
screen "Nas_23" 1280x800
   Softkey "Softkey_F1" at 0,0 size 0x0
      on KeyDown: function_efd93a16()
   IOField "I/O field_6" at 38,288 size 172x31; FormatPattern s999.9; Unit %
      ProcessValue <- "PV"
   IOField "I/O field_1" at 35,197 size 174x31; FormatPattern s999.9; Unit %
      ProcessValue <- "SP"
   IOField "I/O field_2" at 240,288 size 149x31; FormatPattern s999.9; Unit %
      ProcessValue <- "LMN"
   TextField "Text field_8" at 67,259 size 95x25; Text 'Значение'
   TextField "Text field_9" at 75,172 size 84x25; Text 'Задание'
   TextField "Text field_10" at 277,263 size 68x25; Text 'Выход'
   TextField "Text field_11" at 227,174 size 182x25; Text 'Задание в ручном режиме'
   GraphicView "Graphic view_1" at 31,743 size 81x52; Picture "Left_Arrow"
   IOField "I/O field_9" at 253,197 size 156x31; FormatPattern s999.9; Unit Hz
      ProcessValue <- "MAN"
   IOField "I/O field_4" at 543,108 size 163x31; FormatPattern 999.9
      ProcessValue <- "Gain"
   Button "Button_1" at 75,122 size 96x32; TextOff 'Auto / Автомат'
      on Click: ResetBit("Man_ON")
      Appearance <- "Man_ON"
   Button "Button_2" at 277,119 size 96x32; TextOff 'Manual / Ручной'
      on Click: SetBit("Man_ON")
      Appearance <- "Man_ON"
   IOField "I/O field_5" at 544,154 size 163x31; FormatPattern 999999999
      ProcessValue <- "Ti"
   IOField "I/O field_7" at 545,203 size 163x31; FormatPattern 99999
      ProcessValue <- "Td"
   TextField "Text field_4" at 516,112 size 16x25; Text 'P'
   TextField "Text field_5" at 518,158 size 13x25; Text 'I'
   TextField "Text field_6" at 516,207 size 18x25; Text 'D'
   TextField "Text field_3" at 14,6 size 1254x45; Text 'Nasos Xvost №2 / Насос №6'
   Button "Button_5" at 1118,202 size 96x32; TextOff 'Stop / Стоп'
      on Click: ResetBit("06_DB_MOTORS_Nas6_1_OperatorStart")
      Appearance <- "06_DB_MOTORS_Nas6_1_OperatorStart"
   Button "Button_6" at 998,202 size 96x32; TextOff 'Pusk / Пуск'
      Appearance <- "06_DB_MOTORS_Nas6_1_OperatorStart"
      on Click: SetBit("06_DB_MOTORS_Nas6_1_OperatorStart")
   TrendView "Trend view_1" at 17,338 size 1231x398
   IOField "I/O field_3" at 431,289 size 143x31; FormatPattern s999.9; Unit Hz
      ProcessValue <- "PV"
   TextField "Text field_1" at 443,264 size 121x25; Text 'Положение'
   IOField "I/O field_8" at 776,227 size 160x31; Authorization "User administration"; FormatPattern s999.9; Unit Hz
      ProcessValue <- "LMN_HI"
   TextField "Text field_2" at 813,201 size 84x25; Text 'Max'
   IOField "I/O field_10" at 776,292 size 160x31; Authorization "User administration"; FormatPattern s999.9; Unit Hz
      ProcessValue <- "LMN_LO"
   TextField "Text field_7" at 816,267 size 84x25; Text 'Min'
   Circle "Circle_1" at 837,64 size 64x64
      Appearance <- "06_DB_MOTORS_Nas6_1_AnimCodeMotor"
   SymbolicIOField "Символьное поле ввода-вывода_3" at 870,136 size 263x36; TextOn '1'; TextOff '0'; TextList "motor_key"
      Appearance <- "02_DB_DI_BOOL_TVU_neisp"
      ProcessValue <- "Mode_nas_6_1"
   SymbolicIOField "Символьное поле ввода-вывода_1" at 951,79 size 263x36; TextOn '1'; TextOff '0'; TextList "motor_AnimCode"
      ProcessValue <- "06_DB_MOTORS_Nas6_1_AnimCodeMotor"
      Appearance <- "06_DB_MOTORS_Nas6_1_AnimCodeMotor"
   Button "Button_3" at 1152,303 size 80x24; TextOff 'Stop / сброс'
      on Click: SetBit("06_DB_MOTORS_Nas6_1_ResetAlr")
   Softkey "[!Invalid!]Softkey_F1" at 0,0 size 0x0
      on KeyDown: ResetBit("10_DB_PID_7-1р2_Man_ON")
   Softkey "[!Invalid!]Softkey_F3" at 0,0 size 0x0
      on KeyDown: function_b9b71300("10_DB_PID_7-1р2_SP", 1)
   Softkey "[!Invalid!]Softkey_F5" at 0,0 size 0x0
      on KeyDown: function_dd21b452("10_DB_PID_7-1р2_SP", 1)
   Softkey "[!Invalid!]Softkey_F7" at 0,0 size 0x0
      on KeyDown: SetBit("10_DB_PID_7-1р2_Man_ON")
   Softkey "[!Invalid!]Softkey_F9" at 0,0 size 0x0
      on KeyDown: function_b9b71300("10_DB_PID_7-1р2_MAN", 1)
   Softkey "[!Invalid!]Softkey_F11" at 0,0 size 0x0
      on KeyDown: function_dd21b452("10_DB_PID_7-1р2_MAN", 1)
   Softkey "[!Invalid!]Softkey_F2" at 0,0 size 0x0
      on KeyDown: ResetBit("10_DB_PID_7-11р2_Man_ON")
   Softkey "[!Invalid!]Softkey_F4" at 0,0 size 0x0
      on KeyDown: function_b9b71300("10_DB_PID_7-11р2_SP", 1)
   Softkey "[!Invalid!]Softkey_F6" at 0,0 size 0x0
      on KeyDown: function_dd21b452("10_DB_PID_7-11р2_SP", 1)
   Softkey "[!Invalid!]Softkey_F8" at 0,0 size 0x0
      on KeyDown: SetBit("10_DB_PID_7-11р2_Man_ON")
   Softkey "[!Invalid!]Softkey_F10" at 0,0 size 0x0
      on KeyDown: function_b9b71300("10_DB_PID_7-11р2_MAN", 1)
   Softkey "[!Invalid!]Softkey_F12" at 0,0 size 0x0
      on KeyDown: function_dd21b452("10_DB_PID_7-11р2_MAN", 1)

screen "ScreenParametr1" 1280x800
   TextField "Текстовый блок_2" at 0,0 size 1279x39; Text 'Масштабирование аналоговых сигналов 1'
   Group "Group" at 196,40 size 207x56
   Group "Group_1" at 403,40 size 207x56
   Group "Group_2" at 591,40 size 207x56
   Group "Group_4" at 791,40 size 115x56
   Group "Group_5" at 936,40 size 115x56
   Group "Group_3" at 1063,40 size 165x56
   IOField "Поле ввода-вывода_6" at 231,105 size 135x30; FormatPattern s9999.9
      ProcessValue <- "Уставка: MAX"
   IOField "Поле ввода-вывода_1" at 438,105 size 135x30; FormatPattern s999.9
      ProcessValue <- "Уставка: MIN"
   IOField "Поле ввода-вывода_2" at 628,105 size 135x30; FormatPattern s999.9
      ProcessValue <- "Уставка: HH"
   IOField "Поле ввода-вывода_3" at 782,105 size 135x30; FormatPattern s999.9
      ProcessValue <- "Уставка: H"
   IOField "Поле ввода-вывода_4" at 926,105 size 135x30; FormatPattern s999.9
      ProcessValue <- "Уставка: L"
   IOField "Поле ввода-вывода_5" at 1080,105 size 135x30; FormatPattern s999.9
      ProcessValue <- "Уставка: LL"
   IOField "Поле ввода-вывода_13" at 231,181 size 135x30; FormatPattern s9999.9
      ProcessValue <- "Уставка: MAX"
   IOField "Поле ввода-вывода_14" at 438,181 size 135x30; FormatPattern s999.9
      ProcessValue <- "Уставка: MIN"
   IOField "Поле ввода-вывода_15" at 628,181 size 135x30; FormatPattern s999.9
      ProcessValue <- "Уставка: HH"
   IOField "Поле ввода-вывода_16" at 782,181 size 135x30; FormatPattern s999.9
      ProcessValue <- "Уставка: H"
   IOField "Поле ввода-вывода_17" at 926,181 size 135x30; FormatPattern s999.9
      ProcessValue <- "Уставка: L"
   IOField "Поле ввода-вывода_18" at 1080,181 size 135x30; FormatPattern s999.9
      ProcessValue <- "Уставка: LL"
   IOField "Поле ввода-вывода_19" at 231,222 size 135x30; FormatPattern s9999.9
      ProcessValue <- "Уставка: MAX"
   IOField "Поле ввода-вывода_20" at 438,222 size 135x30; FormatPattern s999.9
      ProcessValue <- "Уставка: MIN"
   IOField "Поле ввода-вывода_21" at 628,222 size 135x30; FormatPattern s999.9
      ProcessValue <- "Уставка: HH"
   IOField "Поле ввода-вывода_22" at 782,222 size 135x30; FormatPattern s999.9
      ProcessValue <- "Уставка: H"
   IOField "Поле ввода-вывода_23" at 926,222 size 135x30; FormatPattern s999.9
      ProcessValue <- "Уставка: L"
   IOField "Поле ввода-вывода_24" at 1080,222 size 135x30; FormatPattern s999.9
      ProcessValue <- "Уставка: LL"
   IOField "Поле ввода-вывода_25" at 231,264 size 135x30; FormatPattern s9999.9
      ProcessValue <- "Уставка: MAX"
   IOField "Поле ввода-вывода_26" at 438,264 size 135x30; FormatPattern s999.9
      ProcessValue <- "Уставка: MIN"
   IOField "Поле ввода-вывода_27" at 628,264 size 135x30; FormatPattern s999.9
      ProcessValue <- "Уставка: HH"
   IOField "Поле ввода-вывода_28" at 782,264 size 135x30; FormatPattern s999.9
      ProcessValue <- "Уставка: H"
   IOField "Поле ввода-вывода_29" at 926,264 size 135x30; FormatPattern s999.9
      ProcessValue <- "Уставка: L"
   IOField "Поле ввода-вывода_30" at 1080,264 size 135x30; FormatPattern s999.9
      ProcessValue <- "Уставка: LL"
   IOField "Поле ввода-вывода_31" at 232,304 size 135x30; FormatPattern s9999.9
      ProcessValue <- "Уставка: MAX"
   IOField "Поле ввода-вывода_32" at 439,304 size 135x30; FormatPattern s999.9
      ProcessValue <- "Уставка: MIN"
   IOField "Поле ввода-вывода_33" at 629,304 size 135x30; FormatPattern s999.9
      ProcessValue <- "Уставка: HH"
   IOField "Поле ввода-вывода_34" at 783,304 size 135x30; FormatPattern s999.9
      ProcessValue <- "Уставка: H"
   IOField "Поле ввода-вывода_35" at 927,304 size 135x30; FormatPattern s999.9
      ProcessValue <- "Уставка: L"
   IOField "Поле ввода-вывода_36" at 1081,304 size 135x30; FormatPattern s999.9
      ProcessValue <- "Уставка: LL"
   IOField "Поле ввода-вывода_37" at 232,345 size 135x30; FormatPattern s9999.9
      ProcessValue <- "Уставка: MAX"
   IOField "Поле ввода-вывода_38" at 439,345 size 135x30; FormatPattern s999.9
      ProcessValue <- "Уставка: MIN"
   IOField "Поле ввода-вывода_39" at 629,345 size 135x30; FormatPattern s999.9
      ProcessValue <- "Уставка: HH"
   IOField "Поле ввода-вывода_40" at 783,345 size 135x30; FormatPattern s999.9
      ProcessValue <- "Уставка: H"
   IOField "Поле ввода-вывода_41" at 927,345 size 135x30; FormatPattern s999.9
      ProcessValue <- "Уставка: L"
   IOField "Поле ввода-вывода_42" at 1081,345 size 135x30; FormatPattern s999.9
      ProcessValue <- "Уставка: LL"
   IOField "Поле ввода-вывода_43" at 232,386 size 135x30; FormatPattern s9999.9
      ProcessValue <- "Уставка: MAX"
   IOField "Поле ввода-вывода_44" at 439,386 size 135x30; FormatPattern s999.9
      ProcessValue <- "Уставка: MIN"
   IOField "Поле ввода-вывода_45" at 629,386 size 135x30; FormatPattern s999.9
      ProcessValue <- "Уставка: HH"
   IOField "Поле ввода-вывода_46" at 783,386 size 135x30; FormatPattern s999.9
      ProcessValue <- "Уставка: H"
   IOField "Поле ввода-вывода_47" at 927,386 size 135x30; FormatPattern s999.9
      ProcessValue <- "Уставка: L"
   IOField "Поле ввода-вывода_48" at 1081,386 size 135x30; FormatPattern s999.9
      ProcessValue <- "Уставка: LL"
   IOField "Поле ввода-вывода_49" at 232,428 size 135x30; FormatPattern s9999.9
      ProcessValue <- "Уставка: MAX"
   IOField "Поле ввода-вывода_50" at 439,428 size 135x30; FormatPattern s999.9
      ProcessValue <- "Уставка: MIN"
   IOField "Поле ввода-вывода_51" at 629,428 size 135x30; FormatPattern s999.9
      ProcessValue <- "Уставка: HH"
   IOField "Поле ввода-вывода_52" at 783,428 size 135x30; FormatPattern s999.9
      ProcessValue <- "Уставка: H"
   IOField "Поле ввода-вывода_53" at 927,428 size 135x30; FormatPattern s999.9
      ProcessValue <- "Уставка: L"
   IOField "Поле ввода-вывода_54" at 1081,428 size 135x30; FormatPattern s999.9
      ProcessValue <- "Уставка: LL"
   IOField "Поле ввода-вывода_55" at 232,470 size 135x30; FormatPattern s9999.9
      ProcessValue <- "Уставка: MAX"
   IOField "Поле ввода-вывода_56" at 439,470 size 135x30; FormatPattern s999.9
      ProcessValue <- "Уставка: MIN"
   IOField "Поле ввода-вывода_57" at 629,470 size 135x30; FormatPattern s999.9
      ProcessValue <- "Уставка: HH"
   IOField "Поле ввода-вывода_58" at 783,470 size 135x30; FormatPattern s999.9
      ProcessValue <- "Уставка: H"
   IOField "Поле ввода-вывода_59" at 927,470 size 135x30; FormatPattern s999.9
      ProcessValue <- "Уставка: L"
   IOField "Поле ввода-вывода_60" at 1081,470 size 135x30; FormatPattern s999.9
      ProcessValue <- "Уставка: LL"
   IOField "Поле ввода-вывода_61" at 232,512 size 135x30; FormatPattern s9999.9
      ProcessValue <- "Уставка: MAX"
   IOField "Поле ввода-вывода_62" at 439,512 size 135x30; FormatPattern s999.9
      ProcessValue <- "Уставка: MIN"
   IOField "Поле ввода-вывода_63" at 629,512 size 135x30; FormatPattern s999.9
      ProcessValue <- "Уставка: HH"
   IOField "Поле ввода-вывода_64" at 783,512 size 135x30; FormatPattern s999.9
      ProcessValue <- "Уставка: H"
   IOField "Поле ввода-вывода_65" at 927,512 size 135x30; FormatPattern s999.9
      ProcessValue <- "Уставка: L"
   IOField "Поле ввода-вывода_66" at 1081,512 size 135x30; FormatPattern s999.9
      ProcessValue <- "Уставка: LL"
   IOField "Поле ввода-вывода_67" at 232,551 size 135x30; FormatPattern s9999.9
      ProcessValue <- "Уставка: MAX"
   IOField "Поле ввода-вывода_68" at 439,551 size 135x30; FormatPattern s999.9
      ProcessValue <- "Уставка: MIN"
   IOField "Поле ввода-вывода_69" at 629,551 size 135x30; FormatPattern s999.9
      ProcessValue <- "Уставка: HH"
   IOField "Поле ввода-вывода_70" at 783,551 size 135x30; FormatPattern s999.9
      ProcessValue <- "Уставка: H"
   IOField "Поле ввода-вывода_71" at 927,551 size 135x30; FormatPattern s999.9
      ProcessValue <- "Уставка: L"
   IOField "Поле ввода-вывода_72" at 1081,551 size 135x30; FormatPattern s999.9
      ProcessValue <- "Уставка: LL"
   IOField "Поле ввода-вывода_73" at 232,592 size 135x30; FormatPattern s9999.9
      ProcessValue <- "Уставка: MAX"
   IOField "Поле ввода-вывода_74" at 439,592 size 135x30; FormatPattern s999.9
      ProcessValue <- "Уставка: MIN"
   IOField "Поле ввода-вывода_75" at 629,592 size 135x30; FormatPattern s999.9
      ProcessValue <- "Уставка: HH"
   IOField "Поле ввода-вывода_76" at 783,592 size 135x30; FormatPattern s999.9
      ProcessValue <- "Уставка: H"
   IOField "Поле ввода-вывода_77" at 927,592 size 135x30; FormatPattern s999.9
      ProcessValue <- "Уставка: L"
   IOField "Поле ввода-вывода_78" at 1081,592 size 135x30; FormatPattern s999.9
      ProcessValue <- "Уставка: LL"
   IOField "Поле ввода-вывода_79" at 232,633 size 135x30; FormatPattern s9999.9
      ProcessValue <- "Уставка: MAX"
   IOField "Поле ввода-вывода_80" at 439,633 size 135x30; FormatPattern s999.9
      ProcessValue <- "Уставка: MIN"
   IOField "Поле ввода-вывода_81" at 629,633 size 135x30; FormatPattern s999.9
      ProcessValue <- "Уставка: HH"
   IOField "Поле ввода-вывода_82" at 783,633 size 135x30; FormatPattern s999.9
      ProcessValue <- "Уставка: H"
   IOField "Поле ввода-вывода_83" at 927,633 size 135x30; FormatPattern s999.9
      ProcessValue <- "Уставка: L"
   IOField "Поле ввода-вывода_84" at 1081,633 size 135x30; FormatPattern s999.9
      ProcessValue <- "Уставка: LL"
   IOField "Поле ввода-вывода_85" at 232,673 size 135x30; FormatPattern s9999.9
      ProcessValue <- "Уставка: MAX"
   IOField "Поле ввода-вывода_86" at 439,673 size 135x30; FormatPattern s999.9
      ProcessValue <- "Уставка: MIN"
   IOField "Поле ввода-вывода_87" at 629,673 size 135x30; FormatPattern s999.9
      ProcessValue <- "Уставка: HH"
   IOField "Поле ввода-вывода_88" at 783,673 size 135x30; FormatPattern s999.9
      ProcessValue <- "Уставка: H"
   IOField "Поле ввода-вывода_89" at 927,673 size 135x30; FormatPattern s999.9
      ProcessValue <- "Уставка: L"
   IOField "Поле ввода-вывода_90" at 1081,673 size 135x30; FormatPattern s999.9
      ProcessValue <- "Уставка: LL"
   IOField "Поле ввода-вывода_91" at 232,714 size 135x30; FormatPattern s9999.9
      ProcessValue <- "Уставка: MAX"
   IOField "Поле ввода-вывода_92" at 439,714 size 135x30; FormatPattern s999.9
      ProcessValue <- "Уставка: MIN"
   IOField "Поле ввода-вывода_93" at 629,714 size 135x30; FormatPattern s999.9
      ProcessValue <- "Уставка: HH"
   IOField "Поле ввода-вывода_94" at 783,714 size 135x30; FormatPattern s999.9
      ProcessValue <- "Уставка: H"
   IOField "Поле ввода-вывода_95" at 927,714 size 135x30; FormatPattern s999.9
      ProcessValue <- "Уставка: L"
   IOField "Поле ввода-вывода_96" at 1081,714 size 135x30; FormatPattern s999.9
      ProcessValue <- "Уставка: LL"
   Button "Кнопка_1" at 11,754 size 125x45; TextOff 'Назад'; PictureOff "Left_Arrow"
      on Press: function_efd93a16()
   TextField "Text field_29" at 1104,761 size 175x35; Text 'AI_param2'
   IOField "Поле ввода-вывода_7" at 232,143 size 135x30; FormatPattern s9999.9
      ProcessValue <- "Уставка: MAX"
   IOField "Поле ввода-вывода_8" at 439,143 size 135x30; FormatPattern s999.9
      ProcessValue <- "Уставка: MIN"
   IOField "Поле ввода-вывода_9" at 629,143 size 135x30; FormatPattern s999.9
      ProcessValue <- "Уставка: HH"
   IOField "Поле ввода-вывода_10" at 783,143 size 135x30; FormatPattern s999.9
      ProcessValue <- "Уставка: H"
   IOField "Поле ввода-вывода_11" at 927,143 size 135x30; FormatPattern s999.9
      ProcessValue <- "Уставка: L"
   IOField "Поле ввода-вывода_12" at 1081,143 size 135x30; FormatPattern s999.9
      ProcessValue <- "Уставка: LL"
   TextField "Text field_1" at 216,40 size 165x35; Text 'Инженерный'
   TextField "Text field_2" at 196,61 size 207x35; Text 'верхний диапазон'
   TextField "Text field_3" at 423,40 size 165x35; Text 'Инженерный'
   TextField "Text field_4" at 403,61 size 207x35; Text 'нижний диапазон'
   TextField "Text field_5" at 611,40 size 165x35; Text 'Выше верхняя'
   TextField "Text field_6" at 591,61 size 207x35; Text 'уставка'
   TextField "Text field_9" at 791,40 size 115x35; Text 'Верхняя'
   TextField "Text field_10" at 800,61 size 96x35; Text 'уставка'
   TextField "Text field_11" at 936,40 size 115x35; Text 'Нижняя'
   TextField "Text field_12" at 945,61 size 96x35; Text 'уставка'
   TextField "Text field_7" at 1063,40 size 165x35; Text 'Ниже нижняя'
   TextField "Text field_8" at 1094,61 size 102x35; Text 'уставка'
   Softkey "Softkey_F1" at 0,0 size 0x0
      on KeyDown: function_efd93a16()
   Softkey "Softkey_F10" at 0,0 size 0x0
      on KeyDown: ActivateScreen("ScreenParametr2", 0)

screen "Naraboki" 1280x800
   Button "Кнопка_5" at 11,762 size 125x37; TextOff 'Назад'; PictureOff "Left_Arrow"
      on Press: ActivateScreen("memoscren", 0)
   TextField "Text field_16" at 441,0 size 339x73; Text 'Наработки'
      Appearance <- "Rab_M7"
   IOField "I/O field_1" at 494,145 size 200x51; FormatPattern 99999999
      ProcessValue <- "Hour"
   IOField "I/O field_8" at 700,145 size 66x51; FormatPattern 99
      ProcessValue <- "Minute"
   IOField "I/O field_9" at 773,145 size 66x51; FormatPattern 99
      ProcessValue <- "Second"
   IOField "I/O field_16" at 491,218 size 203x51; FormatPattern 99999999
      ProcessValue <- "Hour"
   IOField "I/O field_17" at 700,218 size 66x51; FormatPattern 99
      ProcessValue <- "Minute"
   IOField "I/O field_18" at 773,219 size 66x51; FormatPattern 99
      ProcessValue <- "Second"
   IOField "I/O field_22" at 494,292 size 200x51; FormatPattern 99999999
      ProcessValue <- "Hour"
   IOField "I/O field_23" at 700,292 size 66x51; FormatPattern 99
      ProcessValue <- "Minute"
   IOField "I/O field_24" at 773,293 size 66x51; FormatPattern 99
      ProcessValue <- "Second"
   IOField "I/O field_25" at 494,366 size 200x51; FormatPattern 99999999
      ProcessValue <- "Hour"
   IOField "I/O field_26" at 700,366 size 66x51; FormatPattern 99
      ProcessValue <- "Minute"
   IOField "I/O field_27" at 773,367 size 66x51; FormatPattern 99
      ProcessValue <- "Second"
   IOField "I/O field_28" at 494,440 size 200x51; FormatPattern 99999999
      ProcessValue <- "Hour"
   IOField "I/O field_29" at 700,440 size 66x51; FormatPattern 99
      ProcessValue <- "Minute"
   IOField "I/O field_30" at 773,441 size 66x51; FormatPattern 99
      ProcessValue <- "Second"
   TextField "Text field_10" at 317,297 size 171x34; Text 'ElectrolyzerWork_1-2 / Насос №3'
   TextField "Text field_11" at 315,149 size 173x34; Text 'ElectrolyzerWork_1-2 / Насос №1'
   TextField "Text field_12" at 317,223 size 171x34; Text 'ElectrolyzerWork_1-2 / Насос №2'
   TextField "Text field_15" at 320,371 size 168x34; Text 'ElectrolyzerWork_1-2 / Насос №4'
   TextField "Text field_17" at 315,445 size 173x34; Text 'ElectrolyzerWork_1-2 / Насос №5'
   IOField "I/O field_40" at 494,514 size 200x51; FormatPattern 99999999
      ProcessValue <- "Hour"
   IOField "I/O field_41" at 700,514 size 66x51; FormatPattern 99
      ProcessValue <- "Minute"
   IOField "I/O field_42" at 773,515 size 66x51; FormatPattern 99
      ProcessValue <- "Second"
   TextField "Text field_18" at 321,519 size 167x34; Text 'ElectrolyzerWork_1-2 / Насос №6'
   TextField "Text field_21" at 527,88 size 77x39; Text 'Hour'
   TextField "Text field_22" at 686,88 size 59x39; Text 'Min'
   TextField "Text field_23" at 762,88 size 55x39; Text 'Sec'
   Button "Кнопка_1" at 1144,760 size 125x37; TextOff 'Назад'; PictureOff "Right_Arrow"
      on Press: ActivateScreen("memoscren", 0)
   Softkey "Softkey_F1" at 0,0 size 0x0
      on KeyDown: function_efd93a16()
   Softkey "Softkey_F10" at 0,0 size 0x0
      on KeyDown: ActivateScreen("Naraboki2", 0)

screen "StartScreen" 1280x800
   Softkey "[!Invalid!]Softkey_F4" at 0,0 size 0x0
      on KeyDown: ActivateScreen("Mill", 0)
   Softkey "[!Invalid!]Softkey_F6" at 0,0 size 0x0
      on KeyDown: ActivateScreen("Oil", 0)
   Softkey "[!Invalid!]Softkey_F8" at 0,0 size 0x0
      on KeyDown: ActivateScreen("Zumpf", 0)
   GraphicView "Graphic view_37" at 1098,144 size 31x29; Picture "Graphic_3"
   GraphicView "Graphic view_38" at 1097,161 size 36x30; Picture "Графика_4"
   GraphicView "Graphic view_29" at 112,653 size 125x83; Picture "Graphic_9"
   GraphicView "Graphic view_33" at 32,586 size 125x83; Picture "Graphic_9"
   GraphicView "Graphic view_4" at 76,199 size 30x30; Picture "Graphic_53"
   GraphicView "Graphic view_2" at 488,89 size 96x72; Picture "gcu"
   GraphicView "Graphic view_21" at 289,269 size 24x23; Picture "Graphic_53"
   GraphicView "Graphic view_26" at 66,268 size 26x25; Picture "Graphic_53"
   GraphicView "Graphic view_19" at 10,199 size 30x30; Picture "Graphic_53"
   GraphicView "Graphic view_1" at 303,234 size 374x277; Picture "MMC_Ch"
   SymbolLibrary "Symbol library_28" at 42,84 size 6x97
   SymbolLibrary "Symbol library_44" at 493,149 size 10x11
   SymbolLibrary "Symbol library_42" at 522,81 size 6x40
   SymbolLibrary "Symbol library_41" at 522,74 size 10x11
   SymbolLibrary "Symbol library_39" at 472,89 size 6x12
   SymbolLibrary "Symbol library_36" at 629,81 size 6x284
   SymbolLibrary "Symbol library_31" at 589,89 size 6x226
   SymbolLibrary "Symbol library_30" at 501,94 size 4x13
   SymbolLibrary "Symbol library_5" at 34,71 size 6x102
   SymbolLibrary "Symbol library_23" at 442,295 size 6x37
   SymbolLibrary "Symbol library_22" at 418,191 size 6x126
   SymbolLibrary "Symbol library_20" at 297,185 size 119x6
   SymbolLibrary "Symbol library_19" at 457,386 size 108x6
   SymbolLibrary "Symbol library_18" at 437,338 size 83x6
   SymbolLibrary "Symbol library_10" at 198,367 size 6x68
   SymbolLibrary "Symbol library_9" at 174,365 size 6x53
   SymbolLibrary "Symbol library_8" at 67,435 size 83x6
   SymbolLibrary "Symbol library_7" at 59,399 size 83x6
   SymbolLibrary "Symbol library_1" at 118,374 size 73x47
      Appearance <- "AnimCodeMotor"
   SymbolLibrary "Symbol library_2" at 517,307 size 93x57
      Appearance <- "AnimCodeMotor"
   SymbolLibrary "Symbol library_3" at 557,355 size 93x57
      Appearance <- "AnimCodeMotor"
   SymbolLibrary "Symbol library_4" at 142,410 size 73x47
      Appearance <- "AnimCodeMotor"
   SymbolLibrary "Symbol library_6" at 174,359 size 10x11
   SymbolLibrary "Symbol library_11" at 193,359 size 11x10
   SymbolLibrary "Symbol library_12" at 180,359 size 17x6
   SymbolLibrary "Symbol library_13" at 186,254 size 6x111
   SymbolLibrary "Symbol library_14" at 181,247 size 11x10
   SymbolLibrary "Symbol library_15" at 104,247 size 79x6
   SymbolLibrary "Symbol library_16" at 97,247 size 10x11
   SymbolLibrary "Symbol library_17" at 97,254 size 6x124
   TextField "Text field_5" at 795,575 size 42x28; Text '6-1 / 36'
   SymbolLibrary "Symbol library_21" at 413,185 size 11x10
   SymbolLibrary "Symbol library_24" at 442,287 size 10x11
   SymbolLibrary "Symbol library_25" at 448,287 size 122x6
   SymbolLibrary "Symbol library_32" at 548,100 size 7x9
   SymbolLibrary "Symbol library_33" at 547,94 size 8x7
   SymbolLibrary "Symbol library_34" at 584,82 size 11x10
   SymbolLibrary "Symbol library_35" at 430,94 size 119x4
   SymbolLibrary "Symbol library_29" at 498,101 size 7x9
   SymbolLibrary "Symbol library_37" at 478,82 size 111x6
   SymbolLibrary "Symbol library_38" at 472,82 size 10x11
   SymbolLibrary "Symbol library_40" at 528,74 size 100x6
   SymbolLibrary "Symbol library_43" at 624,74 size 11x10
   SymbolLibrary "Symbol library_45" at 336,79 size 11x10
   SymbolLibrary "Symbol library_46" at 350,154 size 144x6
   SymbolLibrary "Symbol library_47" at 42,79 size 10x11
   SymbolLibrary "Symbol library_48" at 49,79 size 292x6
   SymbolLibrary "Symbol library_49" at 341,88 size 6x64
   SymbolLibrary "Symbol library_26" at 341,149 size 11x11
   GraphicView "Graphic view_17" at 14,141 size 82x51; Picture "Graphic_38"
   GraphicView "Graphic view_18" at 28,197 size 61x33; Picture "Graphic_41"
   GraphicView "Graphic view_5" at 15,204 size 20x19; Picture "Graphic_52"
   GraphicView "Graphic view_24" at 76,267 size 128x26; Picture "Graphic_41"
   GraphicView "Graphic view_25" at 194,267 size 111x26; Picture "Graphic_41"
   GraphicView "Graphic view_27" at 69,272 size 16x16; Picture "Graphic_52"
   TextField "Text field_3" at 661,580 size 32x18; Text '6-2 / 34'
   Bar "Bar_2" at 649,427 size 174x74; MinimumValue 0; MaximumValue 100
      ProcessValue <- "PV"
   GraphicView "Graphic view_13" at 145,141 size 82x51; Picture "Graphic_38"
   GraphicView "Graphic view_22" at 294,272 size 14x16; Picture "Graphic_52"
   TextField "Text field_2" at 711,436 size 45x26; Text '8-1 / 45'
   TextField "Text field_10" at 30,149 size 29x18; Text '3-2 / 8'
   TextField "Text field_15" at 162,149 size 29x18; Text '3-1 / 9'
   TextField "Text field_16" at 170,249 size 29x18; Text '1-2 / 45'
   TextField "Text field_17" at 139,733 size 51x32; Text '18-2 / 34'
   TextField "Text field_18" at 50,670 size 45x32; Text '18-1 / 23'
   TextField "Text field_20" at 1035,138 size 58x33; Text '9-1 / 5'
   GraphicView "Graphic view_10" at 81,204 size 20x19; Picture "Graphic_52"
   GraphicView "Graphic view_6" at 199,199 size 30x30; Picture "Graphic_53"
   GraphicView "Graphic view_12" at 133,199 size 30x30; Picture "Graphic_53"
   GraphicView "Graphic view_14" at 152,197 size 61x33; Picture "Graphic_41"
   GraphicView "Graphic view_15" at 138,204 size 20x19; Picture "Graphic_52"
   GraphicView "Graphic view_16" at 204,204 size 20x19; Picture "Graphic_52"
   Rectangle "Rectangle_2" at 86,232 size 8x32
      Appearance <- "Rab_ub_trans_3_2"
   Rectangle "Rectangle_3" at 142,232 size 8x32
      Appearance <- "Rab_ub_trans_3_1"
   TextField "Text field_21" at 730,575 size 34x27; Text '6-3 / 35'
   GraphicView "Graphic view_20" at 644,511 size 58x67; Picture "Graphic_57"
   GraphicView "Graphic view_23" at 712,510 size 58x67; Picture "Graphic_57"
   GraphicView "Graphic view_32" at 780,511 size 58x67; Picture "Graphic_57"
   GraphicView "Graphic view_30" at 762,129 size 438x183; Picture "Слой 0 копия_3"
   IOField "I/O field_2" at 861,383 size 83x35; FormatPattern 999.9; Unit %
   IOField "I/O field_3" at 755,383 size 83x35; FormatPattern 999.9; Unit %
   TextField "Text field_27" at 133,439 size 79x36; Text 'Ток 9-1 / Ток 6-2'
   Circle "Circle_2" at 663,535 size 28x28
      Appearance <- "06_DB_MOTORS_Rab_Nas6_2"
   Circle "Circle_3" at 731,534 size 28x28
      Appearance <- "06_DB_MOTORS_Rab_Nas6_3"
   Circle "Circle_4" at 799,535 size 28x28
      Appearance <- "06_DB_MOTORS_Rab_Nas6_1"
   Circle "Circle_7" at 65,147 size 23x23
      Appearance <- "06_DB_MOTORS_Rab_PIT_3_2"
   Circle "Circle_8" at 196,147 size 23x23
      Appearance <- "06_DB_MOTORS_Rab_PIT_3_1"
   IOField "I/O field_6" at 357,266 size 119x35; FormatPattern 999.9; Unit кг/см2
   TextField "Text field_8" at 380,236 size 47x29; Text 'P / Р'
   TextField "Text field_13" at 600,237 size 47x29; Text 'P / Р'
   IOField "I/O field_10" at 30,540 size 75x37; FormatPattern 9999; Unit A
   TextField "Text field_29" at 30,503 size 71x36; Text 'Ток 9-2 / Ток 6-1'
   IOField "I/O field_11" at 635,613 size 71x33; FormatPattern 9999; Unit A
   IOField "I/O field_12" at 715,613 size 65x33; FormatPattern 9999; Unit A
   IOField "I/O field_13" at 786,613 size 67x33; FormatPattern 9999; Unit A
   Circle "Circle_13" at 203,685 size 20x20
      Appearance <- "06_DB_MOTORS_Rab_Nas18_2"
   Circle "Circle_12" at 123,619 size 20x20
      Appearance <- "06_DB_MOTORS_Rab_Nas18_1"
   GraphicView "Graphic view_34" at 272,587 size 125x83; Picture "Graphic_9"
   TextField "Text field_32" at 290,671 size 45x32; Text '13-1 / 45'
   Circle "Circle_15" at 363,620 size 20x20
      Appearance <- "10_DB_Maslonasos_Rabota1"
   TextField "Text field_35" at 720,295 size 34x36; Text '6-1 / 3'
   TextField "Text field_36" at 666,297 size 32x36; Text '6-2 / 1'
   TextField "Text field_37" at 694,299 size 34x31; Text '6-3 / 2'
   TextField "Text field_38" at 21,761 size 77x39; Text '29-7 / ММS'
   TextField "Text field_39" at 148,761 size 83x39; Text '29-7 / Konveer'
   Button "Button_1" at 781,509 size 62x63; TextOff '1'
      on Click: ActivateScreen("Nas_23", 0)
   Button "Button_2" at 711,510 size 62x63; TextOff '1'
      on Click: ActivateScreen("Nas_24", 0)
   Button "Button_3" at 644,510 size 62x63; TextOff '1'
      on Click: ActivateScreen("Nas_25", 0)
   Button "Button_5" at 21,131 size 62x63; TextOff 'Text'
      on Click: ActivateScreen("PIT_3-2", 0)
   Button "Button_6" at 158,134 size 62x63; TextOff 'Text'
      on Click: ActivateScreen("PIT_3-1", 0)
   GraphicView "Graphic view_35" at 569,112 size 96x72; Picture "gcu"
   GraphicView "Graphic view_3" at 955,217 size 41x49; Picture "Graphic_3"
   GraphicView "Graphic view_36" at 954,240 size 46x50; Picture "Графика_4"
   IOField "I/O field_8" at 581,266 size 120x35; FormatPattern 999.9; Unit кг/см2
   IOField "I/O field_5" at 136,484 size 74x37; FormatPattern 9999; Unit A
   SymbolicIOField "Symbolic I/O field_2" at 670,498 size 35x28; TextOff '0'; TextOn '1'; TextList "motor_key1"
      Appearance <- "Mode_nas_6_2"
      ProcessValue <- "Mode_nas_6_2"
   SymbolicIOField "Symbolic I/O field_3" at 741,498 size 35x28; TextOn '1'; TextOff '0'; TextList "motor_key1"
      ProcessValue <- "Mode_nas_6_3"
      Appearance <- "Mode_nas_6_3"
   SymbolicIOField "Symbolic I/O field_4" at 812,498 size 35x28; TextOn '1'; TextOff '0'; TextList "motor_key1"
      Appearance <- "Mode_nas_6_1"
      ProcessValue <- "Mode_nas_6_1"
   TextField "Text field_41" at 252,761 size 118x39; Text '29-7 / Классифик'
   TextField "Text field_42" at 386,761 size 118x39; Text '29-7 / Маслонасос'
   Rectangle "Rectangle_1" at 474,312 size 53x65
      Visibility <- "05_DB_MILL_RABOTA"
   Button "Button_7" at 950,238 size 62x63; TextOff 'Text'
      on Click: ActivateScreen("BAYPAS", 0)
   Button "Button_8" at 1079,127 size 62x63; TextOff 'Text'
      on Click: ActivateScreen("SHIBER", 0)
   Circle "Circle_16" at 262,266 size 32x32
      Appearance <- "07_DB_KONV_RABOTA"
   Circle "Circle_17" at 133,200 size 25x25
      Appearance <- "Rab_ub_trans_3_1"
   Circle "Circle_18" at 79,201 size 25x25
      Appearance <- "Rab_ub_trans_3_2"
   Circle "Circle_20" at 313,320 size 32x32
      Appearance <- "L_telegi"
   DateTimeField "Date/time field_1" at 1026,9 size 236x34
   IOField "I/O field_1" at 293,498 size 74x37; FormatPattern 9999; Unit A
   TextField "Text field_1" at 289,467 size 79x36; Text 'Ток 9-1 / Ток 6-3'
   Softkey "Softkey_F1" at 0,0 size 0x0
      on KeyDown: ActivateScreen("MMS7", 0)
   Softkey "Softkey_F2" at 0,0 size 0x0
      on KeyDown: ActivateScreen("Konv1_2", 0)
   Softkey "Softkey_F3" at 0,0 size 0x0
      on KeyDown: ActivateScreen("klassifikator1", 0)
   Softkey "Softkey_F4" at 0,0 size 0x0
      on KeyDown: ActivateScreen("maslostansiya", 0)

screen "Nas_25" 1280x800
   Softkey "Softkey_F1" at 0,0 size 0x0
      on KeyDown: function_efd93a16()
   IOField "I/O field_6" at 38,288 size 172x31; FormatPattern s999.9; Unit %
      ProcessValue <- "PV"
   IOField "I/O field_1" at 35,197 size 174x31; FormatPattern s999.9; Unit %
      ProcessValue <- "SP"
   IOField "I/O field_2" at 240,288 size 149x31; FormatPattern s999.9; Unit %
      ProcessValue <- "LMN"
   TextField "Text field_8" at 67,259 size 95x25; Text 'Значение'
   TextField "Text field_9" at 75,172 size 84x25; Text 'Задание'
   TextField "Text field_10" at 277,263 size 68x25; Text 'Выход'
   TextField "Text field_11" at 227,174 size 182x25; Text 'Задание в ручном режиме'
   GraphicView "Graphic view_1" at 31,743 size 81x52; Picture "Left_Arrow"
   IOField "I/O field_9" at 253,197 size 156x31; FormatPattern s999.9; Unit Hz
      ProcessValue <- "MAN"
   IOField "I/O field_4" at 543,108 size 163x31; FormatPattern 999.9
      ProcessValue <- "Gain"
   Button "Button_1" at 75,122 size 96x32; TextOff 'Auto / Автомат'
      on Click: ResetBit("Man_ON")
      Appearance <- "Man_ON"
   Button "Button_2" at 277,119 size 96x32; TextOff 'Manual / Ручной'
      on Click: SetBit("Man_ON")
      Appearance <- "Man_ON"
   IOField "I/O field_5" at 544,154 size 163x31; FormatPattern 999999999
      ProcessValue <- "Ti"
   IOField "I/O field_7" at 545,203 size 163x31; FormatPattern 99999
      ProcessValue <- "Td"
   TextField "Text field_4" at 516,112 size 16x25; Text 'P'
   TextField "Text field_5" at 518,158 size 13x25; Text 'I'
   TextField "Text field_6" at 516,207 size 18x25; Text 'D'
   TextField "Text field_3" at 9,9 size 1261x46; Text 'Nasos Xvost №2 / Насос №3'
   Button "Button_5" at 1118,202 size 96x32; TextOff 'Stop / Стоп'
      on Click: ResetBit("06_DB_MOTORS_Nas6_2.OperatorStart")
      Appearance <- "06_DB_MOTORS_Nas6_2.OperatorStart"
   Button "Button_6" at 998,202 size 96x32; TextOff 'Pusk / Пуск'
      on Click: SetBit("06_DB_MOTORS_Nas6_2.OperatorStart")
      Appearance <- "06_DB_MOTORS_Nas6_2.OperatorStart"
   TrendView "Trend view_1" at 17,338 size 1231x398
   IOField "I/O field_3" at 431,289 size 143x31; FormatPattern s999.9; Unit Hz
      ProcessValue <- "PV"
   TextField "Text field_1" at 443,264 size 121x25; Text 'Положение'
   IOField "I/O field_8" at 776,227 size 160x31; Authorization "User administration"; FormatPattern s999.9; Unit Hz
      ProcessValue <- "LMN_HI"
   TextField "Text field_2" at 813,201 size 84x25; Text 'Max'
   IOField "I/O field_10" at 776,292 size 160x31; Authorization "User administration"; FormatPattern s999.9; Unit Hz
      ProcessValue <- "LMN_LO"
   TextField "Text field_7" at 816,267 size 84x25; Text 'Min'
   Circle "Circle_1" at 850,64 size 64x64
      Appearance <- "06_DB_MOTORS_Nas6_2.AnimCodeMotor"
   SymbolicIOField "Символьное поле ввода-вывода_3" at 870,141 size 263x36; TextOn '1'; TextOff '0'; TextList "motor_key"
      Appearance <- "02_DB_DI_BOOL_TVU_neisp"
      ProcessValue <- "Mode_nas_6_2"
   SymbolicIOField "Символьное поле ввода-вывода_1" at 951,79 size 263x36; TextOn '1'; TextOff '0'; TextList "motor_AnimCode"
      ProcessValue <- "06_DB_MOTORS_Nas6_2.AnimCodeMotor"
      Appearance <- "06_DB_MOTORS_Nas6_2.AnimCodeMotor"
   Button "Button_3" at 1152,303 size 80x24; TextOff 'Stop / сброс'
      on Click: SetBit("06_DB_MOTORS_Nas6_2_ResetAlr")
   Softkey "[!Invalid!]Softkey_F1" at 0,0 size 0x0
      on KeyDown: ResetBit("10_DB_PID_7-1р2_Man_ON")
   Softkey "[!Invalid!]Softkey_F3" at 0,0 size 0x0
      on KeyDown: function_b9b71300("10_DB_PID_7-1р2_SP", 1)
   Softkey "[!Invalid!]Softkey_F5" at 0,0 size 0x0
      on KeyDown: function_dd21b452("10_DB_PID_7-1р2_SP", 1)
   Softkey "[!Invalid!]Softkey_F7" at 0,0 size 0x0
      on KeyDown: SetBit("10_DB_PID_7-1р2_Man_ON")
   Softkey "[!Invalid!]Softkey_F9" at 0,0 size 0x0
      on KeyDown: function_b9b71300("10_DB_PID_7-1р2_MAN", 1)
   Softkey "[!Invalid!]Softkey_F11" at 0,0 size 0x0
      on KeyDown: function_dd21b452("10_DB_PID_7-1р2_MAN", 1)
   Softkey "[!Invalid!]Softkey_F2" at 0,0 size 0x0
      on KeyDown: ResetBit("10_DB_PID_7-11р2_Man_ON")
   Softkey "[!Invalid!]Softkey_F4" at 0,0 size 0x0
      on KeyDown: function_b9b71300("10_DB_PID_7-11р2_SP", 1)
   Softkey "[!Invalid!]Softkey_F6" at 0,0 size 0x0
      on KeyDown: function_dd21b452("10_DB_PID_7-11р2_SP", 1)
   Softkey "[!Invalid!]Softkey_F8" at 0,0 size 0x0
      on KeyDown: SetBit("10_DB_PID_7-11р2_Man_ON")
   Softkey "[!Invalid!]Softkey_F10" at 0,0 size 0x0
      on KeyDown: function_b9b71300("10_DB_PID_7-11р2_MAN", 1)
   Softkey "[!Invalid!]Softkey_F12" at 0,0 size 0x0
      on KeyDown: function_dd21b452("10_DB_PID_7-11р2_MAN", 1)

screen "soobshen" 1280x800
   AlarmView "Alarm view_1" at 44,28 size 1213x697
   GraphicView "Graphic view_1" at 31,743 size 81x52; Picture "Left_Arrow"
   Softkey "Softkey_F1" at 0,0 size 0x0
      on KeyDown: function_efd93a16()

screen "Nas_24" 1280x800
   Softkey "Softkey_F1" at 0,0 size 0x0
      on KeyDown: function_efd93a16()
   IOField "I/O field_6" at 38,288 size 172x31; FormatPattern s999.9; Unit %
      ProcessValue <- "PV"
   IOField "I/O field_1" at 35,197 size 174x31; FormatPattern s999.9; Unit %
      ProcessValue <- "SP"
   IOField "I/O field_2" at 240,288 size 149x31; FormatPattern s999.9; Unit %
      ProcessValue <- "LMN"
   TextField "Text field_8" at 67,259 size 95x25; Text 'Значение'
   TextField "Text field_9" at 75,172 size 84x25; Text 'Задание'
   TextField "Text field_10" at 277,263 size 68x25; Text 'Выход'
   TextField "Text field_11" at 227,174 size 182x25; Text 'Задание в ручном режиме'
   GraphicView "Graphic view_1" at 31,743 size 81x52; Picture "Left_Arrow"
   IOField "I/O field_9" at 253,197 size 156x31; FormatPattern s999.9; Unit Hz
      ProcessValue <- "MAN"
   IOField "I/O field_4" at 543,108 size 163x31; FormatPattern 999.9
      ProcessValue <- "Gain"
   Button "Button_1" at 75,122 size 96x32; TextOff 'Auto / Автомат'
      on Click: ResetBit("Man_ON")
      Appearance <- "Man_ON"
   Button "Button_2" at 277,119 size 96x32; TextOff 'Manual / Ручной'
      on Click: SetBit("Man_ON")
      Appearance <- "Man_ON"
   IOField "I/O field_5" at 544,154 size 163x31; FormatPattern 999999999
      ProcessValue <- "Ti"
   IOField "I/O field_7" at 545,203 size 163x31; FormatPattern 99999
      ProcessValue <- "Td"
   TextField "Text field_4" at 516,112 size 16x25; Text 'P'
   TextField "Text field_5" at 518,158 size 13x25; Text 'I'
   TextField "Text field_6" at 516,207 size 18x25; Text 'D'
   TextField "Text field_3" at 9,9 size 1261x46; Text 'Nasos Xvost №2 / Насос №5'
   Button "Button_5" at 1118,202 size 96x32; TextOff 'Stop / Стоп'
      on Click: ResetBit("06_DB_MOTORS_Nas6_3.OperatorStart")
      Appearance <- "06_DB_MOTORS_Nas6_3.OperatorStart"
   Button "Button_6" at 998,202 size 96x32; TextOff 'Pusk / Пуск'
      on Click: SetBit("06_DB_MOTORS_Nas6_3.OperatorStart")
      Appearance <- "06_DB_MOTORS_Nas6_3.OperatorStart"
   TrendView "Trend view_1" at 17,338 size 1231x398
   IOField "I/O field_3" at 431,289 size 143x31; FormatPattern s999.9; Unit Hz
      ProcessValue <- "PV"
   TextField "Text field_1" at 443,264 size 121x25; Text 'Положение'
   IOField "I/O field_8" at 776,227 size 160x31; Authorization "User administration"; FormatPattern s999.9; Unit Hz
      ProcessValue <- "LMN_HI"
   TextField "Text field_2" at 813,201 size 84x25; Text 'Max'
   IOField "I/O field_10" at 776,292 size 160x31; Authorization "User administration"; FormatPattern s999.9; Unit Hz
      ProcessValue <- "LMN_LO"
   TextField "Text field_7" at 816,267 size 84x25; Text 'Min'
   Circle "Circle_1" at 839,73 size 64x64
      Appearance <- "06_DB_MOTORS_Nas6_3_AnimCodeMotor"
   SymbolicIOField "Символьное поле ввода-вывода_3" at 870,145 size 263x36; TextOn '1'; TextOff '0'; TextList "motor_key"
      Appearance <- "02_DB_DI_BOOL_TVU_neisp"
      ProcessValue <- "Mode_nas_6_3"
   SymbolicIOField "Символьное поле ввода-вывода_1" at 951,79 size 263x36; TextOn '1'; TextOff '0'; TextList "motor_AnimCode"
      ProcessValue <- "06_DB_MOTORS_Nas6_3_AnimCodeMotor"
      Appearance <- "06_DB_MOTORS_Nas6_3_AnimCodeMotor"
   Button "Button_3" at 1152,303 size 80x24; TextOff 'Stop / сброс'
      on Click: SetBit("06_DB_MOTORS_Nas6_3_ResetAlr")
   Softkey "[!Invalid!]Softkey_F1" at 0,0 size 0x0
      on KeyDown: ResetBit("10_DB_PID_7-1р2_Man_ON")
   Softkey "[!Invalid!]Softkey_F3" at 0,0 size 0x0
      on KeyDown: function_b9b71300("10_DB_PID_7-1р2_SP", 1)
   Softkey "[!Invalid!]Softkey_F5" at 0,0 size 0x0
      on KeyDown: function_dd21b452("10_DB_PID_7-1р2_SP", 1)
   Softkey "[!Invalid!]Softkey_F7" at 0,0 size 0x0
      on KeyDown: SetBit("10_DB_PID_7-1р2_Man_ON")
   Softkey "[!Invalid!]Softkey_F9" at 0,0 size 0x0
      on KeyDown: function_b9b71300("10_DB_PID_7-1р2_MAN", 1)
   Softkey "[!Invalid!]Softkey_F11" at 0,0 size 0x0
      on KeyDown: function_dd21b452("10_DB_PID_7-1р2_MAN", 1)
   Softkey "[!Invalid!]Softkey_F2" at 0,0 size 0x0
      on KeyDown: ResetBit("10_DB_PID_7-11р2_Man_ON")
   Softkey "[!Invalid!]Softkey_F4" at 0,0 size 0x0
      on KeyDown: function_b9b71300("10_DB_PID_7-11р2_SP", 1)
   Softkey "[!Invalid!]Softkey_F6" at 0,0 size 0x0
      on KeyDown: function_dd21b452("10_DB_PID_7-11р2_SP", 1)
   Softkey "[!Invalid!]Softkey_F8" at 0,0 size 0x0
      on KeyDown: SetBit("10_DB_PID_7-11р2_Man_ON")
   Softkey "[!Invalid!]Softkey_F10" at 0,0 size 0x0
      on KeyDown: function_b9b71300("10_DB_PID_7-11р2_MAN", 1)
   Softkey "[!Invalid!]Softkey_F12" at 0,0 size 0x0
      on KeyDown: function_dd21b452("10_DB_PID_7-11р2_MAN", 1)
*)